// TIA Portal project "EEEB EMBU 4_V17" (V17) (continued)
      ETTSDG4 : Time;   // EFETIVO DO TEMPORIZADOR
      ETTSDG3 : Time;   // EFETIVO DO TEMPORIZADOR
      ETTSDG2 : Time;   // EFETIVO DO TEMPORIZADOR
      ETTSDG1 : Time;   // EFETIVO DO TEMPORIZADOR
   END_VAR
   VAR_TEMP   // added for the SCL form of the ladder/FBD networks
      _w1 : Bool;
   END_VAR
BEGIN

REGION Network 1: Tranforme em segundo o tempo de rodízio dos sopradores
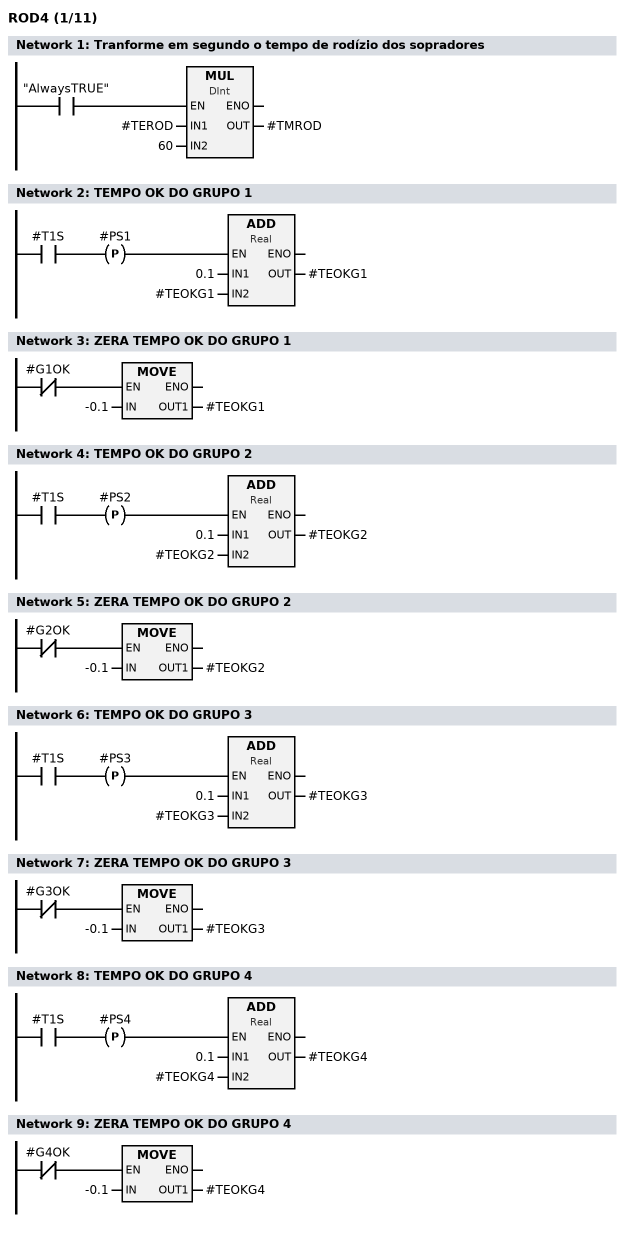
   RUNG wire#powerrail
      Contact( "AlwaysTRUE" )
      { S7_Templates := "SrcType := DInt"; S7_GenerateENO := "TRUE" } Mul(in1 := #TEROD, in2 := 60, out => #TMROD)
   END_RUNG
   // the same network as SCL:
   IF "AlwaysTRUE" THEN #TMROD := #TEROD * 60; END_IF;
END_REGION

REGION Network 2: TEMPO OK DO GRUPO 1
   RUNG wire#powerrail
      Contact( #T1S )
      P_Trig( #PS1 )
      { S7_Templates := "SrcType := Real"; S7_GenerateENO := "TRUE" } Add(in1 := 0.1, in2 := #TEOKG1, out => #TEOKG1)
   END_RUNG
   // the same network as SCL:
   #_w1 := #T1S AND NOT #PS1;   // rising edge
   #PS1 := #T1S;
   IF #_w1 THEN #TEOKG1 := 0.1 + #TEOKG1; END_IF;
END_REGION

REGION Network 3: ZERA TEMPO OK DO GRUPO 1
   RUNG wire#powerrail
      I_Contact( #G1OK )
      { S7_GenerateENO := "TRUE" } Move(in := -0.1, out1 => #TEOKG1)
   END_RUNG
   // the same network as SCL:
   IF NOT #G1OK THEN #TEOKG1 := -0.1; END_IF;
END_REGION

REGION Network 4: TEMPO OK DO GRUPO 2
   RUNG wire#powerrail
      Contact( #T1S )
      P_Trig( #PS2 )
      { S7_Templates := "SrcType := Real"; S7_GenerateENO := "TRUE" } Add(in1 := 0.1, in2 := #TEOKG2, out => #TEOKG2)
   END_RUNG
   // the same network as SCL:
   #_w1 := #T1S AND NOT #PS2;   // rising edge
   #PS2 := #T1S;
   IF #_w1 THEN #TEOKG2 := 0.1 + #TEOKG2; END_IF;
END_REGION

REGION Network 5: ZERA TEMPO OK DO GRUPO 2
   RUNG wire#powerrail
      I_Contact( #G2OK )
      { S7_GenerateENO := "TRUE" } Move(in := -0.1, out1 => #TEOKG2)
   END_RUNG
   // the same network as SCL:
   IF NOT #G2OK THEN #TEOKG2 := -0.1; END_IF;
END_REGION

REGION Network 6: TEMPO OK DO GRUPO 3
   RUNG wire#powerrail
      Contact( #T1S )
      P_Trig( #PS3 )
      { S7_Templates := "SrcType := Real"; S7_GenerateENO := "TRUE" } Add(in1 := 0.1, in2 := #TEOKG3, out => #TEOKG3)
   END_RUNG
   // the same network as SCL:
   #_w1 := #T1S AND NOT #PS3;   // rising edge
   #PS3 := #T1S;
   IF #_w1 THEN #TEOKG3 := 0.1 + #TEOKG3; END_IF;
END_REGION

REGION Network 7: ZERA TEMPO OK DO GRUPO 3
   RUNG wire#powerrail
      I_Contact( #G3OK )
      { S7_GenerateENO := "TRUE" } Move(in := -0.1, out1 => #TEOKG3)
   END_RUNG
   // the same network as SCL:
   IF NOT #G3OK THEN #TEOKG3 := -0.1; END_IF;
END_REGION

REGION Network 8: TEMPO OK DO GRUPO 4
   RUNG wire#powerrail
      Contact( #T1S )
      P_Trig( #PS4 )
      { S7_Templates := "SrcType := Real"; S7_GenerateENO := "TRUE" } Add(in1 := 0.1, in2 := #TEOKG4, out => #TEOKG4)
   END_RUNG
   // the same network as SCL:
   #_w1 := #T1S AND NOT #PS4;   // rising edge
   #PS4 := #T1S;
   IF #_w1 THEN #TEOKG4 := 0.1 + #TEOKG4; END_IF;
END_REGION

REGION Network 9: ZERA TEMPO OK DO GRUPO 4
   RUNG wire#powerrail
      I_Contact( #G4OK )
      { S7_GenerateENO := "TRUE" } Move(in := -0.1, out1 => #TEOKG4)
   END_RUNG
   // the same network as SCL:
   IF NOT #G4OK THEN #TEOKG4 := -0.1; END_IF;
END_REGION

REGION Network 10: DEFINIÇÇÃO DE PRIORIDADE DO GRUPO 1
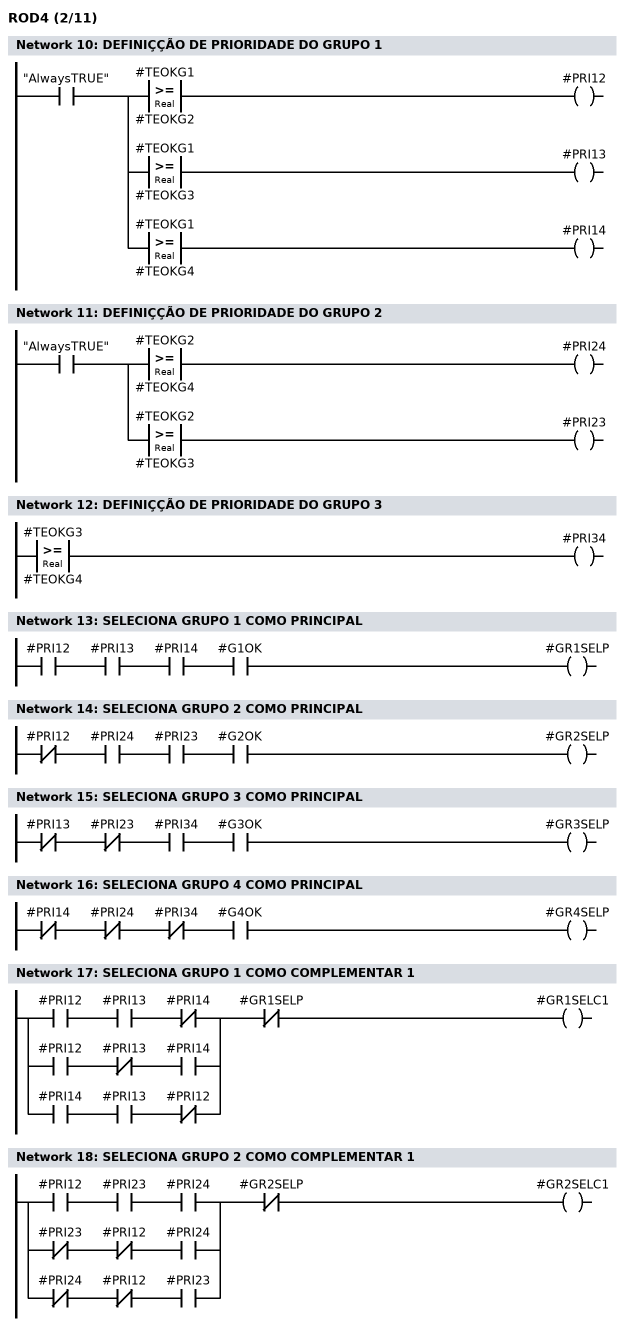
   RUNG wire#powerrail
      Contact( "AlwaysTRUE" )
      wire#w1
      { S7_Templates := "SrcType := Real" } GE_Contact(in1 := #TEOKG1, in2 := #TEOKG2)
      Coil( #PRI12 )
   END_RUNG
   RUNG wire#w1
      { S7_Templates := "SrcType := Real" } GE_Contact(in1 := #TEOKG1, in2 := #TEOKG3)
      Coil( #PRI13 )
   END_RUNG
   RUNG wire#w1
      { S7_Templates := "SrcType := Real" } GE_Contact(in1 := #TEOKG1, in2 := #TEOKG4)
      Coil( #PRI14 )
   END_RUNG
   // the same network as SCL:
   #PRI12 := "AlwaysTRUE" AND (#TEOKG1 >= #TEOKG2);
   #PRI13 := "AlwaysTRUE" AND (#TEOKG1 >= #TEOKG3);
   #PRI14 := "AlwaysTRUE" AND (#TEOKG1 >= #TEOKG4);
END_REGION

REGION Network 11: DEFINIÇÇÃO DE PRIORIDADE DO GRUPO 2
   RUNG wire#powerrail
      Contact( "AlwaysTRUE" )
      wire#w1
      { S7_Templates := "SrcType := Real" } GE_Contact(in1 := #TEOKG2, in2 := #TEOKG4)
      Coil( #PRI24 )
   END_RUNG
   RUNG wire#w1
      { S7_Templates := "SrcType := Real" } GE_Contact(in1 := #TEOKG2, in2 := #TEOKG3)
      Coil( #PRI23 )
   END_RUNG
   // the same network as SCL:
   #PRI24 := "AlwaysTRUE" AND (#TEOKG2 >= #TEOKG4);
   #PRI23 := "AlwaysTRUE" AND (#TEOKG2 >= #TEOKG3);
END_REGION

REGION Network 12: DEFINIÇÇÃO DE PRIORIDADE DO GRUPO 3
   RUNG wire#powerrail
      { S7_Templates := "SrcType := Real" } GE_Contact(in1 := #TEOKG3, in2 := #TEOKG4)
      Coil( #PRI34 )
   END_RUNG
   // the same network as SCL:
   #PRI34 := #TEOKG3 >= #TEOKG4;
END_REGION

REGION Network 13: SELECIONA GRUPO 1 COMO PRINCIPAL
   RUNG wire#powerrail
      Contact( #PRI12 )
      Contact( #PRI13 )
      Contact( #PRI14 )
      Contact( #G1OK )
      Coil( #GR1SELP )
   END_RUNG
   // the same network as SCL:
   #GR1SELP := #PRI12 AND #PRI13 AND #PRI14 AND #G1OK;
END_REGION

REGION Network 14: SELECIONA GRUPO 2 COMO PRINCIPAL
   RUNG wire#powerrail
      I_Contact( #PRI12 )
      Contact( #PRI24 )
      Contact( #PRI23 )
      Contact( #G2OK )
      Coil( #GR2SELP )
   END_RUNG
   // the same network as SCL:
   #GR2SELP := NOT #PRI12 AND #PRI24 AND #PRI23 AND #G2OK;
END_REGION

REGION Network 15: SELECIONA GRUPO 3 COMO PRINCIPAL
   RUNG wire#powerrail
      I_Contact( #PRI13 )
      I_Contact( #PRI23 )
      Contact( #PRI34 )
      Contact( #G3OK )
      Coil( #GR3SELP )
   END_RUNG
   // the same network as SCL:
   #GR3SELP := NOT #PRI13 AND NOT #PRI23 AND #PRI34 AND #G3OK;
END_REGION

REGION Network 16: SELECIONA GRUPO 4 COMO PRINCIPAL
   RUNG wire#powerrail
      I_Contact( #PRI14 )
      I_Contact( #PRI24 )
      I_Contact( #PRI34 )
      Contact( #G4OK )
      Coil( #GR4SELP )
   END_RUNG
   // the same network as SCL:
   #GR4SELP := NOT #PRI14 AND NOT #PRI24 AND NOT #PRI34 AND #G4OK;
END_REGION

REGION Network 17: SELECIONA GRUPO 1 COMO COMPLEMENTAR 1
   RUNG wire#powerrail
      Contact( #PRI12 )
      Contact( #PRI13 )
      I_Contact( #PRI14 )
      wire#w1
      I_Contact( #GR1SELP )
      Coil( #GR1SELC1 )
   END_RUNG
   RUNG wire#powerrail
      Contact( #PRI12 )
      I_Contact( #PRI13 )
      Contact( #PRI14 )
   END_RUNG wire#w1
   RUNG wire#powerrail
      Contact( #PRI14 )
      Contact( #PRI13 )
      I_Contact( #PRI12 )
   END_RUNG wire#w1
   // the same network as SCL:
   #GR1SELC1 := ((#PRI12 AND #PRI13 AND NOT #PRI14) OR (#PRI12 AND NOT #PRI13 AND #PRI14) OR (#PRI14 AND #PRI13 AND NOT #PRI12)) AND NOT #GR1SELP;
END_REGION

REGION Network 18: SELECIONA GRUPO 2 COMO COMPLEMENTAR 1
   RUNG wire#powerrail
      Contact( #PRI12 )
      Contact( #PRI23 )
      Contact( #PRI24 )
      wire#w1
      I_Contact( #GR2SELP )
      Coil( #GR2SELC1 )
   END_RUNG
   RUNG wire#powerrail
      I_Contact( #PRI23 )
      I_Contact( #PRI12 )
      Contact( #PRI24 )
   END_RUNG wire#w1
   RUNG wire#powerrail
      I_Contact( #PRI24 )
      I_Contact( #PRI12 )
      Contact( #PRI23 )
   END_RUNG wire#w1
   // the same network as SCL:
   #GR2SELC1 := ((#PRI12 AND #PRI23 AND #PRI24) OR (NOT #PRI23 AND NOT #PRI12 AND #PRI24) OR (NOT #PRI24 AND NOT #PRI12 AND #PRI23)) AND NOT #GR2SELP;
END_REGION

REGION Network 19: SELECIONA GRUPO 3 COMO COMPLEMENTAR 1
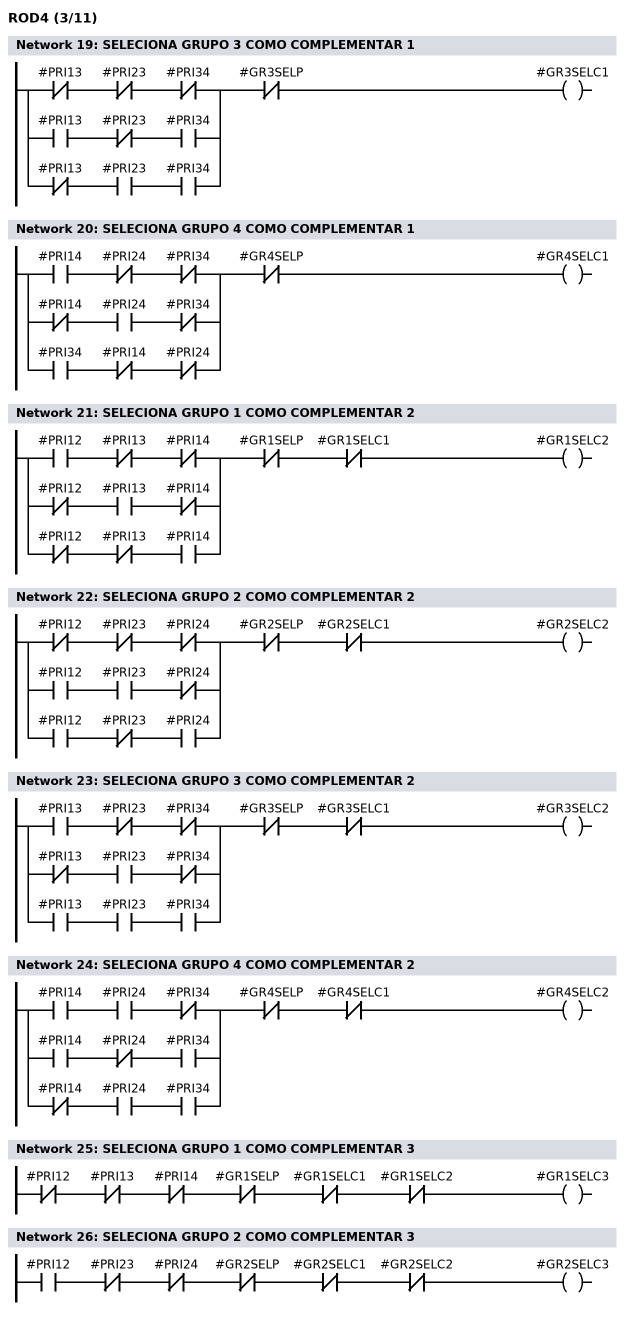
   RUNG wire#powerrail
      I_Contact( #PRI13 )
      I_Contact( #PRI23 )
      I_Contact( #PRI34 )
      wire#w1
      I_Contact( #GR3SELP )
      Coil( #GR3SELC1 )
   END_RUNG
   RUNG wire#powerrail
      Contact( #PRI13 )
      I_Contact( #PRI23 )
      Contact( #PRI34 )
   END_RUNG wire#w1
   RUNG wire#powerrail
      I_Contact( #PRI13 )
      Contact( #PRI23 )
      Contact( #PRI34 )
   END_RUNG wire#w1
   // the same network as SCL:
   #GR3SELC1 := ((NOT #PRI13 AND NOT #PRI23 AND NOT #PRI34) OR (#PRI13 AND NOT #PRI23 AND #PRI34) OR (NOT #PRI13 AND #PRI23 AND #PRI34)) AND NOT #GR3SELP;
END_REGION

REGION Network 20: SELECIONA GRUPO 4 COMO COMPLEMENTAR 1
   RUNG wire#powerrail
      Contact( #PRI14 )
      I_Contact( #PRI24 )
      I_Contact( #PRI34 )
      wire#w1
      I_Contact( #GR4SELP )
      Coil( #GR4SELC1 )
   END_RUNG
   RUNG wire#powerrail
      I_Contact( #PRI14 )
      Contact( #PRI24 )
      I_Contact( #PRI34 )
   END_RUNG wire#w1
   RUNG wire#powerrail
      Contact( #PRI34 )
      I_Contact( #PRI14 )
      I_Contact( #PRI24 )
   END_RUNG wire#w1
   // the same network as SCL:
   #GR4SELC1 := ((#PRI14 AND NOT #PRI24 AND NOT #PRI34) OR (NOT #PRI14 AND #PRI24 AND NOT #PRI34) OR (#PRI34 AND NOT #PRI14 AND NOT #PRI24)) AND NOT #GR4SELP;
END_REGION

REGION Network 21: SELECIONA GRUPO 1 COMO COMPLEMENTAR 2
   RUNG wire#powerrail
      Contact( #PRI12 )
      I_Contact( #PRI13 )
      I_Contact( #PRI14 )
      wire#w1
      I_Contact( #GR1SELP )
      I_Contact( #GR1SELC1 )
      Coil( #GR1SELC2 )
   END_RUNG
   RUNG wire#powerrail
      I_Contact( #PRI12 )
      Contact( #PRI13 )
      I_Contact( #PRI14 )
   END_RUNG wire#w1
   RUNG wire#powerrail
      I_Contact( #PRI12 )
      I_Contact( #PRI13 )
      Contact( #PRI14 )
   END_RUNG wire#w1
   // the same network as SCL:
   #GR1SELC2 := ((#PRI12 AND NOT #PRI13 AND NOT #PRI14) OR (NOT #PRI12 AND #PRI13 AND NOT #PRI14) OR (NOT #PRI12 AND NOT #PRI13 AND #PRI14)) AND NOT #GR1SELP AND NOT #GR1SELC1;
END_REGION

REGION Network 22: SELECIONA GRUPO 2 COMO COMPLEMENTAR 2
   RUNG wire#powerrail
      I_Contact( #PRI12 )
      I_Contact( #PRI23 )
      I_Contact( #PRI24 )
      wire#w1
      I_Contact( #GR2SELP )
      I_Contact( #GR2SELC1 )
      Coil( #GR2SELC2 )
   END_RUNG
   RUNG wire#powerrail
      Contact( #PRI12 )
      Contact( #PRI23 )
      I_Contact( #PRI24 )
   END_RUNG wire#w1
   RUNG wire#powerrail
      Contact( #PRI12 )
      I_Contact( #PRI23 )
      Contact( #PRI24 )
   END_RUNG wire#w1
   // the same network as SCL:
   #GR2SELC2 := ((NOT #PRI12 AND NOT #PRI23 AND NOT #PRI24) OR (#PRI12 AND #PRI23 AND NOT #PRI24) OR (#PRI12 AND NOT #PRI23 AND #PRI24)) AND NOT #GR2SELP AND NOT #GR2SELC1;
END_REGION

REGION Network 23: SELECIONA GRUPO 3 COMO COMPLEMENTAR 2
   RUNG wire#powerrail
      Contact( #PRI13 )
      I_Contact( #PRI23 )
      I_Contact( #PRI34 )
      wire#w1
      I_Contact( #GR3SELP )
      I_Contact( #GR3SELC1 )
      Coil( #GR3SELC2 )
   END_RUNG
   RUNG wire#powerrail
      I_Contact( #PRI13 )
      Contact( #PRI23 )
      I_Contact( #PRI34 )
   END_RUNG wire#w1
   RUNG wire#powerrail
      Contact( #PRI13 )
      Contact( #PRI23 )
      Contact( #PRI34 )
   END_RUNG wire#w1
   // the same network as SCL:
   #GR3SELC2 := ((#PRI13 AND NOT #PRI23 AND NOT #PRI34) OR (NOT #PRI13 AND #PRI23 AND NOT #PRI34) OR (#PRI13 AND #PRI23 AND #PRI34)) AND NOT #GR3SELP AND NOT #GR3SELC1;
END_REGION

REGION Network 24: SELECIONA GRUPO 4 COMO COMPLEMENTAR 2
   RUNG wire#powerrail
      Contact( #PRI14 )
      Contact( #PRI24 )
      I_Contact( #PRI34 )
      wire#w1
      I_Contact( #GR4SELP )
      I_Contact( #GR4SELC1 )
      Coil( #GR4SELC2 )
   END_RUNG
   RUNG wire#powerrail
      Contact( #PRI14 )
      I_Contact( #PRI24 )
      Contact( #PRI34 )
   END_RUNG wire#w1
   RUNG wire#powerrail
      I_Contact( #PRI14 )
      Contact( #PRI24 )
      Contact( #PRI34 )
   END_RUNG wire#w1
   // the same network as SCL:
   #GR4SELC2 := ((#PRI14 AND #PRI24 AND NOT #PRI34) OR (#PRI14 AND NOT #PRI24 AND #PRI34) OR (NOT #PRI14 AND #PRI24 AND #PRI34)) AND NOT #GR4SELP AND NOT #GR4SELC1;
END_REGION

REGION Network 25: SELECIONA GRUPO 1 COMO COMPLEMENTAR 3
   RUNG wire#powerrail
      I_Contact( #PRI12 )
      I_Contact( #PRI13 )
      I_Contact( #PRI14 )
      I_Contact( #GR1SELP )
      I_Contact( #GR1SELC1 )
      I_Contact( #GR1SELC2 )
      Coil( #GR1SELC3 )
   END_RUNG
   // the same network as SCL:
   #GR1SELC3 := NOT #PRI12 AND NOT #PRI13 AND NOT #PRI14 AND NOT #GR1SELP AND NOT #GR1SELC1 AND NOT #GR1SELC2;
END_REGION

REGION Network 26: SELECIONA GRUPO 2 COMO COMPLEMENTAR 3
   RUNG wire#powerrail
      Contact( #PRI12 )
      I_Contact( #PRI23 )
      I_Contact( #PRI24 )
      I_Contact( #GR2SELP )
      I_Contact( #GR2SELC1 )
      I_Contact( #GR2SELC2 )
      Coil( #GR2SELC3 )
   END_RUNG
   // the same network as SCL:
   #GR2SELC3 := #PRI12 AND NOT #PRI23 AND NOT #PRI24 AND NOT #GR2SELP AND NOT #GR2SELC1 AND NOT #GR2SELC2;
END_REGION

REGION Network 27: SELECIONA GRUPO 3 COMO COMPLEMENTAR 3
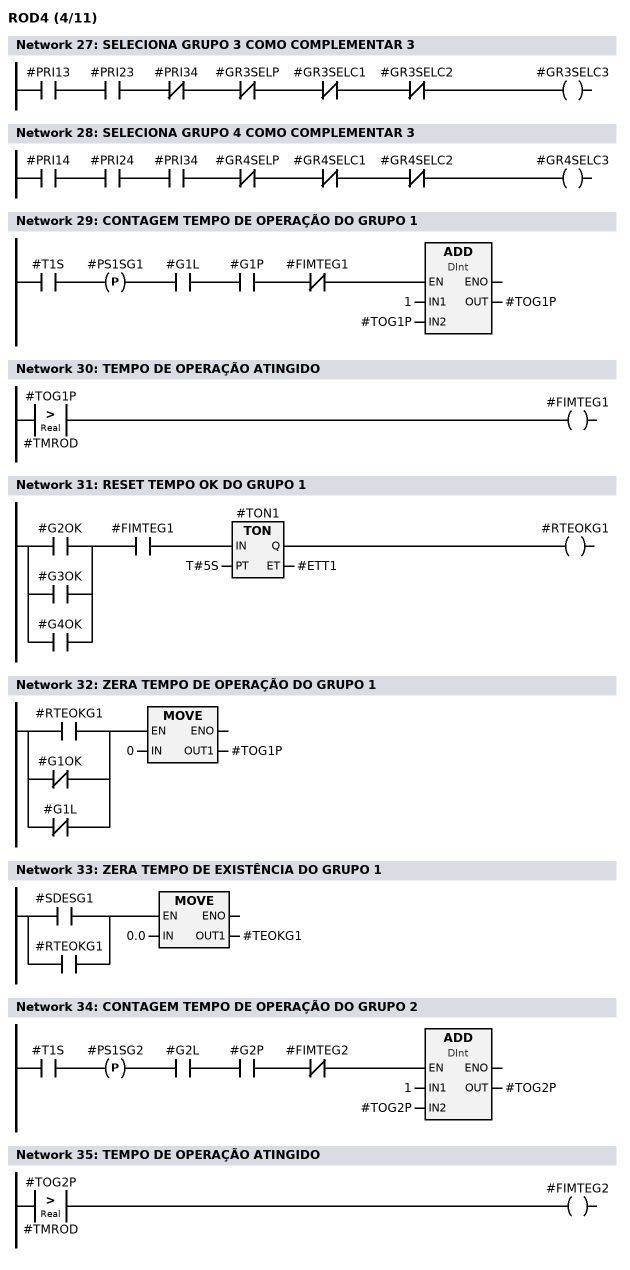
   RUNG wire#powerrail
      Contact( #PRI13 )
      Contact( #PRI23 )
      I_Contact( #PRI34 )
      I_Contact( #GR3SELP )
      I_Contact( #GR3SELC1 )
      I_Contact( #GR3SELC2 )
      Coil( #GR3SELC3 )
   END_RUNG
   // the same network as SCL:
   #GR3SELC3 := #PRI13 AND #PRI23 AND NOT #PRI34 AND NOT #GR3SELP AND NOT #GR3SELC1 AND NOT #GR3SELC2;
END_REGION

REGION Network 28: SELECIONA GRUPO 4 COMO COMPLEMENTAR 3
   RUNG wire#powerrail
      Contact( #PRI14 )
      Contact( #PRI24 )
      Contact( #PRI34 )
      I_Contact( #GR4SELP )
      I_Contact( #GR4SELC1 )
      I_Contact( #GR4SELC2 )
      Coil( #GR4SELC3 )
   END_RUNG
   // the same network as SCL:
   #GR4SELC3 := #PRI14 AND #PRI24 AND #PRI34 AND NOT #GR4SELP AND NOT #GR4SELC1 AND NOT #GR4SELC2;
END_REGION

REGION Network 29: CONTAGEM TEMPO DE OPERAÇÃO DO GRUPO 1
   RUNG wire#powerrail
      Contact( #T1S )
      P_Trig( #PS1SG1 )
      Contact( #G1L )
      Contact( #G1P )
      I_Contact( #FIMTEG1 )
      { S7_Templates := "SrcType := DInt"; S7_GenerateENO := "TRUE" } Add(in1 := 1, in2 := #TOG1P, out => #TOG1P)
   END_RUNG
   // the same network as SCL:
   #_w1 := #T1S AND NOT #PS1SG1;   // rising edge
   #PS1SG1 := #T1S;
   IF #_w1 AND #G1L AND #G1P AND NOT #FIMTEG1 THEN #TOG1P := 1 + #TOG1P; END_IF;
END_REGION

REGION Network 30: TEMPO DE OPERAÇÃO ATINGIDO
   RUNG wire#powerrail
      { S7_Templates := "SrcType := Real" } GT_Contact(in1 := #TOG1P, in2 := #TMROD)
      Coil( #FIMTEG1 )
   END_RUNG
   // the same network as SCL:
   #FIMTEG1 := #TOG1P > #TMROD;
END_REGION

REGION Network 31: RESET TEMPO OK DO GRUPO 1
   #TON1(IN := (#G2OK OR #G3OK OR #G4OK) AND #FIMTEG1, PT := T#5S, ET => #ETT1);   // TON
   #RTEOKG1 := #TON1.Q;
END_REGION

REGION Network 32: ZERA TEMPO DE OPERAÇÃO DO GRUPO 1
   RUNG wire#powerrail
      Contact( #RTEOKG1 )
      wire#w1
      { S7_GenerateENO := "TRUE" } Move(in := 0, out1 => #TOG1P)
   END_RUNG
   RUNG wire#powerrail
      I_Contact( #G1OK )
   END_RUNG wire#w1
   RUNG wire#powerrail
      I_Contact( #G1L )
   END_RUNG wire#w1
   // the same network as SCL:
   IF #RTEOKG1 OR NOT #G1OK OR NOT #G1L THEN #TOG1P := 0; END_IF;
END_REGION

REGION Network 33: ZERA TEMPO DE EXISTÊNCIA DO GRUPO 1
   RUNG wire#powerrail
      Contact( #SDESG1 )
      wire#w1
      { S7_GenerateENO := "TRUE" } Move(in := 0.0, out1 => #TEOKG1)
   END_RUNG
   RUNG wire#powerrail
      Contact( #RTEOKG1 )
   END_RUNG wire#w1
   // the same network as SCL:
   IF #SDESG1 OR #RTEOKG1 THEN #TEOKG1 := 0.0; END_IF;
END_REGION

REGION Network 34: CONTAGEM TEMPO DE OPERAÇÃO DO GRUPO 2
   RUNG wire#powerrail
      Contact( #T1S )
      P_Trig( #PS1SG2 )
      Contact( #G2L )
      Contact( #G2P )
      I_Contact( #FIMTEG2 )
      { S7_Templates := "SrcType := DInt"; S7_GenerateENO := "TRUE" } Add(in1 := 1, in2 := #TOG2P, out => #TOG2P)
   END_RUNG
   // the same network as SCL:
   #_w1 := #T1S AND NOT #PS1SG2;   // rising edge
   #PS1SG2 := #T1S;
   IF #_w1 AND #G2L AND #G2P AND NOT #FIMTEG2 THEN #TOG2P := 1 + #TOG2P; END_IF;
END_REGION

REGION Network 35: TEMPO DE OPERAÇÃO ATINGIDO
   RUNG wire#powerrail
      { S7_Templates := "SrcType := Real" } GT_Contact(in1 := #TOG2P, in2 := #TMROD)
      Coil( #FIMTEG2 )
   END_RUNG
   // the same network as SCL:
   #FIMTEG2 := #TOG2P > #TMROD;
END_REGION

REGION Network 36: RESET TEMPO OK DO GRUPO 2
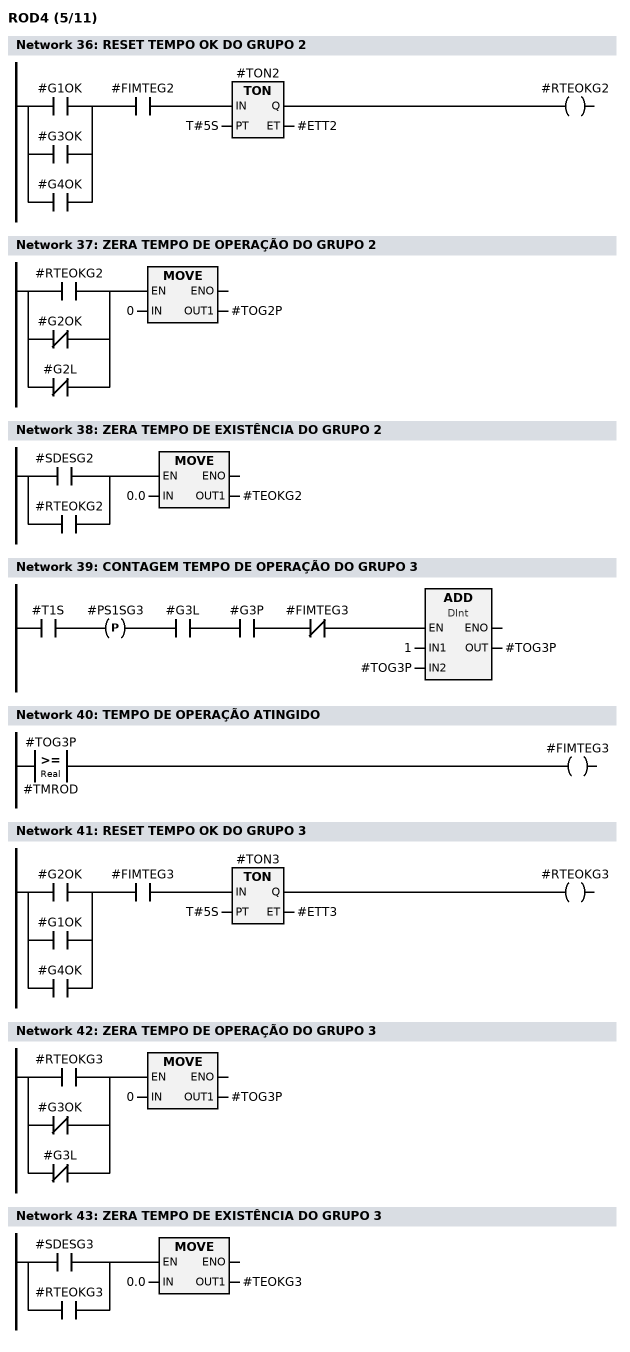
   #TON2(IN := (#G1OK OR #G3OK OR #G4OK) AND #FIMTEG2, PT := T#5S, ET => #ETT2);   // TON
   #RTEOKG2 := #TON2.Q;
END_REGION

REGION Network 37: ZERA TEMPO DE OPERAÇÃO DO GRUPO 2
   RUNG wire#powerrail
      Contact( #RTEOKG2 )
      wire#w1
      { S7_GenerateENO := "TRUE" } Move(in := 0, out1 => #TOG2P)
   END_RUNG
   RUNG wire#powerrail
      I_Contact( #G2OK )
   END_RUNG wire#w1
   RUNG wire#powerrail
      I_Contact( #G2L )
   END_RUNG wire#w1
   // the same network as SCL:
   IF #RTEOKG2 OR NOT #G2OK OR NOT #G2L THEN #TOG2P := 0; END_IF;
END_REGION

REGION Network 38: ZERA TEMPO DE EXISTÊNCIA DO GRUPO 2
   RUNG wire#powerrail
      Contact( #SDESG2 )
      wire#w1
      { S7_GenerateENO := "TRUE" } Move(in := 0.0, out1 => #TEOKG2)
   END_RUNG
   RUNG wire#powerrail
      Contact( #RTEOKG2 )
   END_RUNG wire#w1
   // the same network as SCL:
   IF #SDESG2 OR #RTEOKG2 THEN #TEOKG2 := 0.0; END_IF;
END_REGION

REGION Network 39: CONTAGEM TEMPO DE OPERAÇÃO DO GRUPO 3
   RUNG wire#powerrail
      Contact( #T1S )
      P_Trig( #PS1SG3 )
      Contact( #G3L )
      Contact( #G3P )
      I_Contact( #FIMTEG3 )
      { S7_Templates := "SrcType := DInt"; S7_GenerateENO := "TRUE" } Add(in1 := 1, in2 := #TOG3P, out => #TOG3P)
   END_RUNG
   // the same network as SCL:
   #_w1 := #T1S AND NOT #PS1SG3;   // rising edge
   #PS1SG3 := #T1S;
   IF #_w1 AND #G3L AND #G3P AND NOT #FIMTEG3 THEN #TOG3P := 1 + #TOG3P; END_IF;
END_REGION

REGION Network 40: TEMPO DE OPERAÇÃO ATINGIDO
   RUNG wire#powerrail
      { S7_Templates := "SrcType := Real" } GE_Contact(in1 := #TOG3P, in2 := #TMROD)
      Coil( #FIMTEG3 )
   END_RUNG
   // the same network as SCL:
   #FIMTEG3 := #TOG3P >= #TMROD;
END_REGION

REGION Network 41: RESET TEMPO OK DO GRUPO 3
   #TON3(IN := (#G2OK OR #G1OK OR #G4OK) AND #FIMTEG3, PT := T#5S, ET => #ETT3);   // TON
   #RTEOKG3 := #TON3.Q;
END_REGION

REGION Network 42: ZERA TEMPO DE OPERAÇÃO DO GRUPO 3
   RUNG wire#powerrail
      Contact( #RTEOKG3 )
      wire#w1
      { S7_GenerateENO := "TRUE" } Move(in := 0, out1 => #TOG3P)
   END_RUNG
   RUNG wire#powerrail
      I_Contact( #G3OK )
   END_RUNG wire#w1
   RUNG wire#powerrail
      I_Contact( #G3L )
   END_RUNG wire#w1
   // the same network as SCL:
   IF #RTEOKG3 OR NOT #G3OK OR NOT #G3L THEN #TOG3P := 0; END_IF;
END_REGION

REGION Network 43: ZERA TEMPO DE EXISTÊNCIA DO GRUPO 3
   RUNG wire#powerrail
      Contact( #SDESG3 )
      wire#w1
      { S7_GenerateENO := "TRUE" } Move(in := 0.0, out1 => #TEOKG3)
   END_RUNG
   RUNG wire#powerrail
      Contact( #RTEOKG3 )
   END_RUNG wire#w1
   // the same network as SCL:
   IF #SDESG3 OR #RTEOKG3 THEN #TEOKG3 := 0.0; END_IF;
END_REGION

REGION Network 44: CONTAGEM TEMPO DE OPERAÇÃO DO GRUPO 4
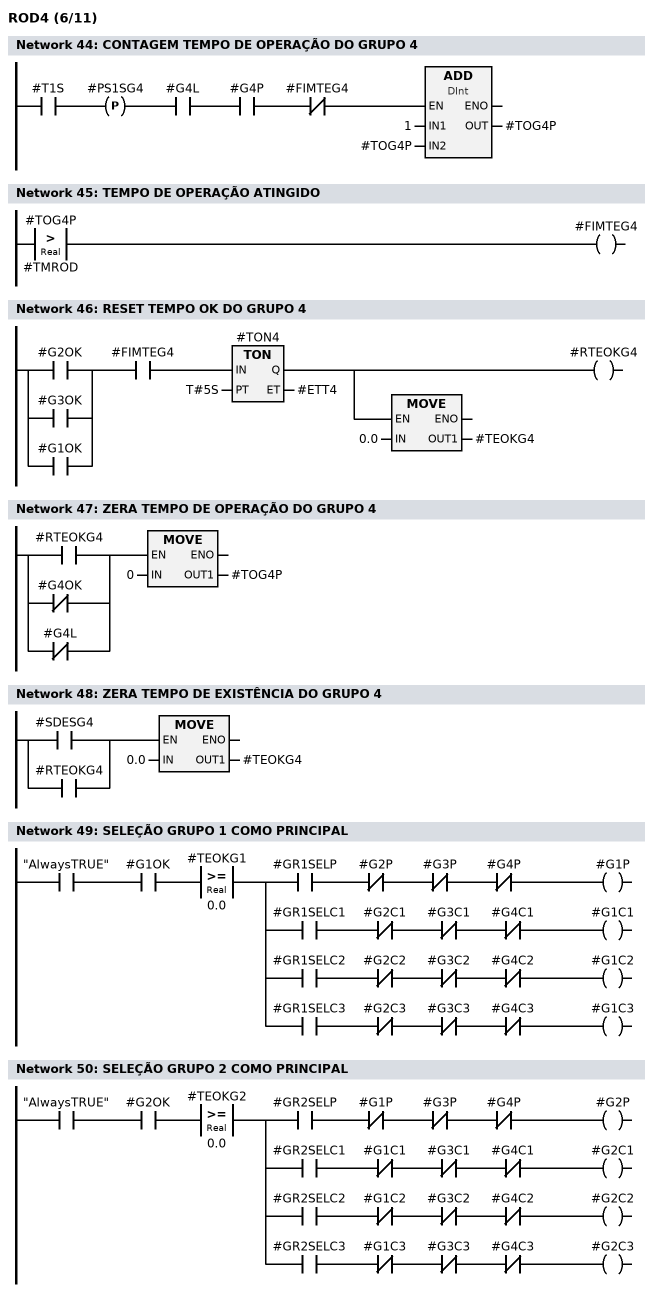
   RUNG wire#powerrail
      Contact( #T1S )
      P_Trig( #PS1SG4 )
      Contact( #G4L )
      Contact( #G4P )
      I_Contact( #FIMTEG4 )
      { S7_Templates := "SrcType := DInt"; S7_GenerateENO := "TRUE" } Add(in1 := 1, in2 := #TOG4P, out => #TOG4P)
   END_RUNG
   // the same network as SCL:
   #_w1 := #T1S AND NOT #PS1SG4;   // rising edge
   #PS1SG4 := #T1S;
   IF #_w1 AND #G4L AND #G4P AND NOT #FIMTEG4 THEN #TOG4P := 1 + #TOG4P; END_IF;
END_REGION

REGION Network 45: TEMPO DE OPERAÇÃO ATINGIDO
   RUNG wire#powerrail
      { S7_Templates := "SrcType := Real" } GT_Contact(in1 := #TOG4P, in2 := #TMROD)
      Coil( #FIMTEG4 )
   END_RUNG
   // the same network as SCL:
   #FIMTEG4 := #TOG4P > #TMROD;
END_REGION

REGION Network 46: RESET TEMPO OK DO GRUPO 4
   #TON4(IN := (#G2OK OR #G3OK OR #G1OK) AND #FIMTEG4, PT := T#5S, ET => #ETT4);   // TON
   #RTEOKG4 := #TON4.Q;
   IF #TON4.Q THEN #TEOKG4 := 0.0; END_IF;
END_REGION

REGION Network 47: ZERA TEMPO DE OPERAÇÃO DO GRUPO 4
   RUNG wire#powerrail
      Contact( #RTEOKG4 )
      wire#w1
      { S7_GenerateENO := "TRUE" } Move(in := 0, out1 => #TOG4P)
   END_RUNG
   RUNG wire#powerrail
      I_Contact( #G4OK )
   END_RUNG wire#w1
   RUNG wire#powerrail
      I_Contact( #G4L )
   END_RUNG wire#w1
   // the same network as SCL:
   IF #RTEOKG4 OR NOT #G4OK OR NOT #G4L THEN #TOG4P := 0; END_IF;
END_REGION

REGION Network 48: ZERA TEMPO DE EXISTÊNCIA DO GRUPO 4
   RUNG wire#powerrail
      Contact( #SDESG4 )
      wire#w1
      { S7_GenerateENO := "TRUE" } Move(in := 0.0, out1 => #TEOKG4)
   END_RUNG
   RUNG wire#powerrail
      Contact( #RTEOKG4 )
   END_RUNG wire#w1
   // the same network as SCL:
   IF #SDESG4 OR #RTEOKG4 THEN #TEOKG4 := 0.0; END_IF;
END_REGION

REGION Network 49: SELEÇÃO GRUPO 1 COMO PRINCIPAL
   RUNG wire#powerrail
      Contact( "AlwaysTRUE" )
      Contact( #G1OK )
      { S7_Templates := "SrcType := Real" } GE_Contact(in1 := #TEOKG1, in2 := 0.0)
      wire#w1
      Contact( #GR1SELP )
      I_Contact( #G2P )
      I_Contact( #G3P )
      I_Contact( #G4P )
      Coil( #G1P )
   END_RUNG
   RUNG wire#w1
      Contact( #GR1SELC1 )
      I_Contact( #G2C1 )
      I_Contact( #G3C1 )
      I_Contact( #G4C1 )
      Coil( #G1C1 )
   END_RUNG
   RUNG wire#w1
      Contact( #GR1SELC2 )
      I_Contact( #G2C2 )
      I_Contact( #G3C2 )
      I_Contact( #G4C2 )
      Coil( #G1C2 )
   END_RUNG
   RUNG wire#w1
      Contact( #GR1SELC3 )
      I_Contact( #G2C3 )
      I_Contact( #G3C3 )
      I_Contact( #G4C3 )
      Coil( #G1C3 )
   END_RUNG
   // the same network as SCL:
   #_w1 := "AlwaysTRUE" AND #G1OK AND (#TEOKG1 >= 0.0);
   #G1P := #_w1 AND #GR1SELP AND NOT #G2P AND NOT #G3P AND NOT #G4P;
   #G1C1 := #_w1 AND #GR1SELC1 AND NOT #G2C1 AND NOT #G3C1 AND NOT #G4C1;
   #G1C2 := #_w1 AND #GR1SELC2 AND NOT #G2C2 AND NOT #G3C2 AND NOT #G4C2;
   #G1C3 := #_w1 AND #GR1SELC3 AND NOT #G2C3 AND NOT #G3C3 AND NOT #G4C3;
END_REGION

REGION Network 50: SELEÇÃO GRUPO 2 COMO PRINCIPAL
   RUNG wire#powerrail
      Contact( "AlwaysTRUE" )
      Contact( #G2OK )
      { S7_Templates := "SrcType := Real" } GE_Contact(in1 := #TEOKG2, in2 := 0.0)
      wire#w1
      Contact( #GR2SELP )
      I_Contact( #G1P )
      I_Contact( #G3P )
      I_Contact( #G4P )
      Coil( #G2P )
   END_RUNG
   RUNG wire#w1
      Contact( #GR2SELC1 )
      I_Contact( #G1C1 )
      I_Contact( #G3C1 )
      I_Contact( #G4C1 )
      Coil( #G2C1 )
   END_RUNG
   RUNG wire#w1
      Contact( #GR2SELC2 )
      I_Contact( #G1C2 )
      I_Contact( #G3C2 )
      I_Contact( #G4C2 )
      Coil( #G2C2 )
   END_RUNG
   RUNG wire#w1
      Contact( #GR2SELC3 )
      I_Contact( #G1C3 )
      I_Contact( #G3C3 )
      I_Contact( #G4C3 )
      Coil( #G2C3 )
   END_RUNG
   // the same network as SCL:
   #_w1 := "AlwaysTRUE" AND #G2OK AND (#TEOKG2 >= 0.0);
   #G2P := #_w1 AND #GR2SELP AND NOT #G1P AND NOT #G3P AND NOT #G4P;
   #G2C1 := #_w1 AND #GR2SELC1 AND NOT #G1C1 AND NOT #G3C1 AND NOT #G4C1;
   #G2C2 := #_w1 AND #GR2SELC2 AND NOT #G1C2 AND NOT #G3C2 AND NOT #G4C2;
   #G2C3 := #_w1 AND #GR2SELC3 AND NOT #G1C3 AND NOT #G3C3 AND NOT #G4C3;
END_REGION

REGION Network 51: SELEÇÃO GRUPO 3 COMO PRINCIPAL
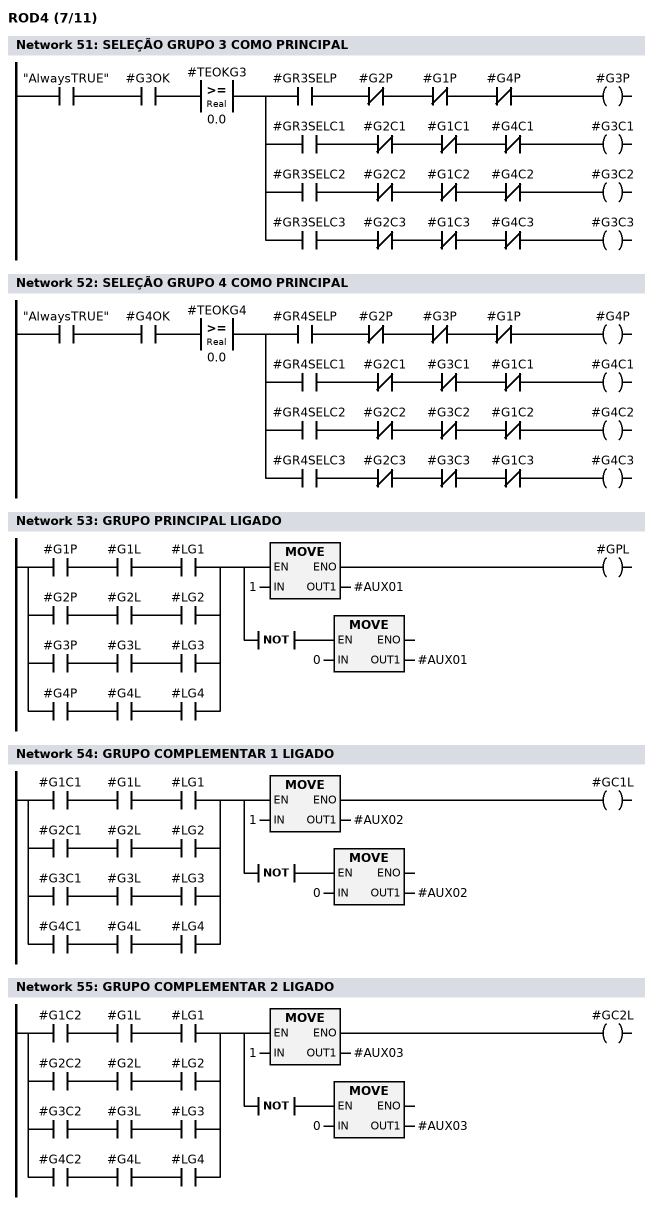
   RUNG wire#powerrail
      Contact( "AlwaysTRUE" )
      Contact( #G3OK )
      { S7_Templates := "SrcType := Real" } GE_Contact(in1 := #TEOKG3, in2 := 0.0)
      wire#w1
      Contact( #GR3SELP )
      I_Contact( #G2P )
      I_Contact( #G1P )
      I_Contact( #G4P )
      Coil( #G3P )
   END_RUNG
   RUNG wire#w1
      Contact( #GR3SELC1 )
      I_Contact( #G2C1 )
      I_Contact( #G1C1 )
      I_Contact( #G4C1 )
      Coil( #G3C1 )
   END_RUNG
   RUNG wire#w1
      Contact( #GR3SELC2 )
      I_Contact( #G2C2 )
      I_Contact( #G1C2 )
      I_Contact( #G4C2 )
      Coil( #G3C2 )
   END_RUNG
   RUNG wire#w1
      Contact( #GR3SELC3 )
      I_Contact( #G2C3 )
      I_Contact( #G1C3 )
      I_Contact( #G4C3 )
      Coil( #G3C3 )
   END_RUNG
   // the same network as SCL:
   #_w1 := "AlwaysTRUE" AND #G3OK AND (#TEOKG3 >= 0.0);
   #G3P := #_w1 AND #GR3SELP AND NOT #G2P AND NOT #G1P AND NOT #G4P;
   #G3C1 := #_w1 AND #GR3SELC1 AND NOT #G2C1 AND NOT #G1C1 AND NOT #G4C1;
   #G3C2 := #_w1 AND #GR3SELC2 AND NOT #G2C2 AND NOT #G1C2 AND NOT #G4C2;
   #G3C3 := #_w1 AND #GR3SELC3 AND NOT #G2C3 AND NOT #G1C3 AND NOT #G4C3;
END_REGION

REGION Network 52: SELEÇÃO GRUPO 4 COMO PRINCIPAL
   RUNG wire#powerrail
      Contact( "AlwaysTRUE" )
      Contact( #G4OK )
      { S7_Templates := "SrcType := Real" } GE_Contact(in1 := #TEOKG4, in2 := 0.0)
      wire#w1
      Contact( #GR4SELP )
      I_Contact( #G2P )
      I_Contact( #G3P )
      I_Contact( #G1P )
      Coil( #G4P )
   END_RUNG
   RUNG wire#w1
      Contact( #GR4SELC1 )
      I_Contact( #G2C1 )
      I_Contact( #G3C1 )
      I_Contact( #G1C1 )
      Coil( #G4C1 )
   END_RUNG
   RUNG wire#w1
      Contact( #GR4SELC2 )
      I_Contact( #G2C2 )
      I_Contact( #G3C2 )
      I_Contact( #G1C2 )
      Coil( #G4C2 )
   END_RUNG
   RUNG wire#w1
      Contact( #GR4SELC3 )
      I_Contact( #G2C3 )
      I_Contact( #G3C3 )
      I_Contact( #G1C3 )
      Coil( #G4C3 )
   END_RUNG
   // the same network as SCL:
   #_w1 := "AlwaysTRUE" AND #G4OK AND (#TEOKG4 >= 0.0);
   #G4P := #_w1 AND #GR4SELP AND NOT #G2P AND NOT #G3P AND NOT #G1P;
   #G4C1 := #_w1 AND #GR4SELC1 AND NOT #G2C1 AND NOT #G3C1 AND NOT #G1C1;
   #G4C2 := #_w1 AND #GR4SELC2 AND NOT #G2C2 AND NOT #G3C2 AND NOT #G1C2;
   #G4C3 := #_w1 AND #GR4SELC3 AND NOT #G2C3 AND NOT #G3C3 AND NOT #G1C3;
END_REGION

REGION Network 53: GRUPO PRINCIPAL LIGADO
   RUNG wire#powerrail
      Contact( #G1P )
      Contact( #G1L )
      Contact( #LG1 )
      wire#w1
      { S7_GenerateENO := "TRUE" } Move(in := 1, out1 => #AUX01)
      Coil( #GPL )
   END_RUNG
   RUNG wire#powerrail
      Contact( #G2P )
      Contact( #G2L )
      Contact( #LG2 )
   END_RUNG wire#w1
   RUNG wire#powerrail
      Contact( #G3P )
      Contact( #G3L )
      Contact( #LG3 )
   END_RUNG wire#w1
   RUNG wire#powerrail
      Contact( #G4P )
      Contact( #G4L )
      Contact( #LG4 )
   END_RUNG wire#w1
   RUNG wire#w1
      Not()
      { S7_GenerateENO := "TRUE" } Move(in := 0, out1 => #AUX01)
   END_RUNG
   // the same network as SCL:
   // ENO of a box is taken as its EN; it also drops when the box reports an error
   #_w1 := (#G1P AND #G1L AND #LG1) OR (#G2P AND #G2L AND #LG2) OR (#G3P AND #G3L AND #LG3) OR (#G4P AND #G4L AND #LG4);
   IF #_w1 THEN #AUX01 := 1; END_IF;
   #GPL := #_w1;
   IF NOT #_w1 THEN #AUX01 := 0; END_IF;
END_REGION

REGION Network 54: GRUPO COMPLEMENTAR 1 LIGADO
   RUNG wire#powerrail
      Contact( #G1C1 )
      Contact( #G1L )
      Contact( #LG1 )
      wire#w1
      { S7_GenerateENO := "TRUE" } Move(in := 1, out1 => #AUX02)
      Coil( #GC1L )
   END_RUNG
   RUNG wire#powerrail
      Contact( #G2C1 )
      Contact( #G2L )
      Contact( #LG2 )
   END_RUNG wire#w1
   RUNG wire#powerrail
      Contact( #G3C1 )
      Contact( #G3L )
      Contact( #LG3 )
   END_RUNG wire#w1
   RUNG wire#powerrail
      Contact( #G4C1 )
      Contact( #G4L )
      Contact( #LG4 )
   END_RUNG wire#w1
   RUNG wire#w1
      Not()
      { S7_GenerateENO := "TRUE" } Move(in := 0, out1 => #AUX02)
   END_RUNG
   // the same network as SCL:
   // ENO of a box is taken as its EN; it also drops when the box reports an error
   #_w1 := (#G1C1 AND #G1L AND #LG1) OR (#G2C1 AND #G2L AND #LG2) OR (#G3C1 AND #G3L AND #LG3) OR (#G4C1 AND #G4L AND #LG4);
   IF #_w1 THEN #AUX02 := 1; END_IF;
   #GC1L := #_w1;
   IF NOT #_w1 THEN #AUX02 := 0; END_IF;
END_REGION

